
Template "01_One_Nav_Level" 1920x1080
   Gauge "gaugeDiagStateUpdate" at 566,2 size 50x50; CaptionText 'SIMATIC'
      on Change: "CheckDiagState"()
      ProcessValue <- "@DiagnosticsIndicatorTag"
   TextField "txtTitleBar" at 8,11 size 361x32; Text 'Application Name / Applikation / 江苏睿博环保再生胶系统'
   GraphicView "gfxNavigationIcon" at 1879,15 size 23x19; Picture "Hamburger_Icon"
   Button "btnNavigation" at 1862,0 size 56x48; TextOff 'Text'
      on Click: function_cf6f4242("GraphX_Slidein_Right", 1)
   TextField "模板_文本域_1" at 283,78 size 160x19; Text '全胎粉'
   TextField "txtTitleBar_1" at 12,1031 size 62x32; Text 'Application Name / Applikation / 冷水:'
   TextField "txtTitleBar_2" at 173,1031 size 62x32; Text 'Application Name / Applikation / 热水:'
   TextField "txtTitleBar_3" at 345,1031 size 62x32; Text 'Application Name / Applikation / 备料:'
   TextField "txtTitleBar_4" at 1752,1030 size 69x32; Text 'Application Name / Applikation / 数据库:'
   TextField "txtTitleBar_5" at 1587,1031 size 69x32; Text 'Application Name / Applikation / 云数据:'
   AlarmView "模板_报警视图_1" at 495,1024 size 1069x52
   IOField "I/O 域_58" at 1096,73 size 129x32; FormatPattern 999999.9; Unit  H
   IOField "I/O 域_59" at 1406,75 size 130x32; FormatPattern 99999999.9; Unit  Kg
   ScreenModuleView "HMI_Indicator_Square_1" at 1834,1033 size 28x28; ScreenModuleType ""
      Guid_{11997190-149293} <- "数据库字符串_Connect_CND"
      Guid_{11997190-149297} <- "数据库字符串_Query_Error"
      Guid_{11997190-149295} <- "数据库字符串_Query_Done"
   ScreenModuleView "HMI_Indicator_Square_2" at 1669,1033 size 28x28; ScreenModuleType ""
      Guid_{11997190-149295} <- "数据库字符串_Query_Done"
      Guid_{11997190-149293} <- "数据库字符串_Connect_CND"
      Guid_{11997190-149297} <- "数据库字符串_Query_Error"
   TextField "模板_文本域_2" at 77,80 size 73x19; Text '请选择'
   Button "btnStartscreen" at 1,2 size 411x45; TextOff 'Text'
      on Click: "ActivateStartScreen"()
   TextField "txtStateHeadline" at 75,55 size 123x23; Text 'State / Status / 运行配方'
   TextField "txtRecipeHeadline" at 281,55 size 154x23; Text 'Current Recipe / Rezeptur / 运行模式'
   TextField "txtOperatorHeadline" at 527,55 size 129x23; Text 'Operator / Bediener / 当前用户'
   IOField "ioOperator" at 527,72 size 126x30; FormatPattern ??????????????????
      ProcessValue <- "CurrentUserName"
   Button "btnState" at 202,56 size 40x40; TextOff '...'; PictureOff "More_Icon"
      on Click: "ShowRecipePopUp"()
   Button "btnRecipe" at 449,56 size 40x40; TextOff '...'; PictureOff "More_Icon"
   Rectangle "rectState" at 0,48 size 56x56
      Appearance <- "CurrentMachineState"
   GraphicIOField "gioDiagState" at 1874,60 size 32x32; PictureList "DiagState_3"
      ProcessValue <- "DiagState"
   Button "btnDiagState" at 1862,48 size 56x56; TextOff 'Text'
   Button "btnOperator" at 669,56 size 40x40; TextOff '...'; PictureOff "More_Icon"
      on Click: function_efd93a16("Template_Logon", 800, 300, -1, -1, 1)
   TextField "txtOperatorHeadline_1" at 768,55 size 129x23; Text 'Date and Time / Bediener / 当前时间'
   Button "btnOperator_1" at 995,56 size 40x40; TextOff '...'; PictureOff "More_Icon"
   DateTimeField "Template_Date/time field_1" at 768,72 size 208x30
   IOField "ioOperator_1" at 69,1033 size 99x30; FormatPattern 99.9; Unit m³/h
   IOField "ioOperator_2" at 230,1033 size 97x30; FormatPattern 99.9; Unit m³/h
   IOField "ioOperator_3" at 402,1033 size 72x30; FormatPattern 99.9; Unit %
   TextField "txtOperatorHeadline_2" at 1094,57 size 129x23; Text 'Date and Time / Bediener / 累计运行时间'
   Button "btnOperator_2" at 1321,58 size 40x40; TextOff '...'; PictureOff "More_Icon"
   TextField "txtOperatorHeadline_3" at 1403,58 size 129x23; Text 'Date and Time / Bediener / 累计产量'
   Button "btnOperator_3" at 1630,59 size 40x40; TextOff '...'; PictureOff "More_Icon"

PopupScreen "Template_Logon" 320x352
   on ClearScreen: ResetBit("PopUpBackground")
   on GenerateScreen: SetBit("PopUpBackground")
   TextField "Template_Text field_1" at 16,0 size 215x40; Text 'Login / 登录'
   Button "Button_2" at 16,240 size 288x40; TextOn 'LOGIN / ANMELDEN / 登录'; TextOff 'LOGIN / ANMELDEN / 登录'
      on Click: function_a9b89908("Password", "UserName"); function_efd93a16("Template_Logon", 0, 0, 0, -1, 1)
   IOField "I/O field_1" at 16,84 size 288x40; FormatPattern ??????????????????????????????
      ProcessValue <- "UserName"
   TextField "Text field_1" at 16,56 size 288x24; Text 'User Name / Name / 用户名'
   IOField "I/O field_2" at 16,168 size 288x40; FormatPattern ??????????????????????????????
      ProcessValue <- "Password"
   TextField "Text field_2" at 16,140 size 288x24; Text 'Password / Passwort / 密码'
   Button "Button_1" at 16,296 size 288x40; TextOn 'CLOSE / SCHLIESSEN / 取消'; TextOff 'CLOSE / SCHLIESSEN / 取消'
      on Click: function_efd93a16("Template_Logon", 0, 0, 0, -1, 1)
      on Press: function_b14e0dd5("ButtonDown", 0)
      Appearance <- "ButtonDown"

PopupScreen "Template_Logon_Logoff" 320x352
   on ClearScreen: ResetBit("PopUpBackground")
   on GenerateScreen: SetBit("PopUpBackground")
   TextField "Template_Text field_1" at 16,0 size 215x40; Text 'Login'
   Button "Button_2" at 16,240 size 136x40; TextOn 'LOG OFF / ABMELDEN'; TextOff 'LOG OFF / ABMELDEN'
      on Click: function_f23ef4c9()
   IOField "I/O field_1" at 16,84 size 288x40; FormatPattern ??????????????????????????????
      ProcessValue <- "UserName"
   TextField "Text field_1" at 16,56 size 288x24; Text 'User Name / Name'
   IOField "I/O field_2" at 16,168 size 288x40; FormatPattern ??????????????????????????????
      ProcessValue <- "Password"
   TextField "Text field_2" at 16,140 size 288x24; Text 'Password / Passwort'
   Button "Button_1" at 16,296 size 288x40; TextOn 'CLOSE / SCHLIESSEN'; TextOff 'CLOSE / SCHLIESSEN'
      on Click: function_efd93a16("Template_Logon_Logoff", 0, 0, 0, -1, 1)
      on Press: function_b14e0dd5("ButtonDown", 0)
      Appearance <- "ButtonDown"
   Button "Button_3" at 168,240 size 136x40; TextOn 'LOGIN / ANMELDEN'; TextOff 'LOGIN / ANMELDEN'
      on Click: function_a9b89908("Password", "UserName"); function_efd93a16("Template_Logon_Logoff", 0, 0, 0, -1, 1)

PopupScreen "Template_Operating_Mode" 424x360
   on ClearScreen: ResetBit("PopUpBackground")
   on GenerateScreen: SetBit("PopUpBackground")
   TextField "Template_Text field_1" at 14,0 size 336x40; Text 'Operating Mode / Betriebsmodus / 单螺杆操作'
   Button "Button_2" at 352,66 size 40x40; TextOff 'Text'; PictureOff "More_Icon"; PictureOn "More_Icon"
      on Click: function_efd93a16("Template_Operating_Mode", 0, 0, 0, -1, 1)
   Button "Button_3" at 352,130 size 40x40; TextOff 'Text'; PictureOff "More_Icon"; PictureOn "More_Icon"
      on Click: function_efd93a16("Template_Operating_Mode", 0, 0, 0, -1, 1)
   Button "Button_4" at 352,189 size 40x40; TextOff 'Text'; PictureOff "More_Icon"; PictureOn "More_Icon"
   Button "Button_1" at 352,254 size 40x40; TextOff 'Text'; PictureOff "More_Icon"; PictureOn "More_Icon"
   TextField "txtParameter7_3" at 32,63 size 163x24; Text 'Demo Mode / Current Mode / 演示模式'
   TextField "txtParameter7_5" at 31,89 size 319x24; Text 'Current Mode / 通过控制台仿真数据给触摸屏进行系统演示'
   TextField "txtParameter7_1" at 32,129 size 163x24; Text 'Test Mode / Current Mode / 测试模式'
   TextField "txtParameter7_2" at 31,155 size 319x24; Text 'Current Mode / 通过控制台仿真数据给触摸屏进行系统演示'

PopupScreen "Template_Recipe" 700x420
   on ClearScreen: ResetBit("PopUpBackground")
   on GenerateScreen: SetBit("PopUpBackground")
   TextField "Template_Text field_1" at 14,0 size 500x40; Text 'Recipe / Rezeptur'
   Button "Button_1" at 220,364 size 260x40; TextOn 'CLOSE / SCHLIESSEN'; TextOff 'CLOSE / SCHLIESSEN / 确定'
      on Click: function_efd93a16("Template_Recipe", 0, 0, 0, -1, 1)
      on Press: function_b14e0dd5("ButtonDown", 0)
      Appearance <- "ButtonDown"

PopupScreen "OptionPanel_4_Buttons_1" 390x648
   Button "btnCloseOptionPanel" at 0,0 size 40x648; TextOff 'CLOSE'; PictureOff "Jog_Forward"
      on Press: function_efd93a16("OptionPanel_4_Buttons_1", 0, 0, 0, 2, 2)
   TextField "txtOptionPanel" at 108,16 size 260x40; Text 'Option Panel Title / Titel Option Panel'
   Button "btnOption1" at 80,72 size 240x40; TextOff 'Option 1 / Move to Home Position'
   Button "btnOption2" at 80,128 size 240x40; TextOff 'Option 2 / Move to Home Position'
   Button "btnOption3" at 80,184 size 240x40; TextOff 'Option 3 / RESET'
   Button "btnOption4" at 80,240 size 240x40; TextOff 'Option 4 / RESET'
   GraphicView "gvOptionPanel" at 80,30 size 18x12; Picture "ManFunctions_Off"

PopupScreen "OptionPanel_4_Buttons" 390x648
   Button "btnCloseOptionPanel" at 0,0 size 40x648; TextOff 'CLOSE'; PictureOff "Jog_Forward"
      on Press: function_efd93a16("OptionPanel_4_Buttons", 0, 0, 0, 2, 2)
   TextField "txtOptionPanel" at 108,16 size 260x40; Text 'Option Panel Title / Titel Option Panel'
   Button "btnOption1" at 80,72 size 240x40; TextOff 'Option 1 / Move to Home Position'
   Button "btnOption2" at 80,128 size 240x40; TextOff 'Option 2 / Move to Home Position'
   Button "btnOption3" at 80,184 size 240x40; TextOff 'Option 3 / RESET'
   Button "btnOption4" at 80,240 size 240x40; TextOff 'Option 4 / RESET'
   GraphicView "gvOptionPanel" at 80,30 size 18x12; Picture "ManFunctions_Off"

PopupScreen "OptionPanel_4_Large_Buttons" 390x648
   Button "btnCloseOptionPanel" at 0,0 size 40x648; TextOff 'CLOSE'; PictureOff "Jog_Forward"
      on Press: function_efd93a16("OptionPanel_4_Large_Buttons", 0, 0, 0, 2, 2)
   TextField "txtOptionPanel" at 108,16 size 260x40; Text 'Option Panel Title / Titel Option Panel'
   GraphicView "gvOptionPanel" at 80,30 size 18x12; Picture "ManFunctions_Off"
   Button "btnOption1" at 80,72 size 112x96; TextOff 'Option 1 / Move to Home Position'
   Button "btnOption2" at 208,72 size 112x96; TextOff 'Option 2 / Move to Home Position'
   Button "btnOption3" at 80,184 size 112x96; TextOff 'Option 3 / Move to Home Position'
   Button "btnOption4" at 208,184 size 112x96; TextOff 'Option 4 / Move to Home Position'

PopupScreen "OptionPanel_8_Buttons" 390x648
   Button "btnCloseOptionPanel" at 0,0 size 40x648; TextOff 'CLOSE'; PictureOff "Jog_Forward"
      on Press: function_efd93a16("OptionPanel_8_Buttons", 0, 0, 0, 2, 2)
   TextField "txtOptionPanel" at 108,16 size 260x40; Text 'Option Panel Title / Titel Option Panel'
   GraphicView "gvOptionPanel" at 80,30 size 18x12; Picture "ManFunctions_Off"
   Button "btnOption1" at 80,72 size 112x40; TextOff 'Option 1 / Move to Home Position'
   Button "btnOption2" at 208,72 size 112x40; TextOff 'Option 2 / Move to Home Position'
   Button "btnOption3" at 80,128 size 112x40; TextOff 'Option 3 / Move to Home Position'
   Button "btnOption4" at 208,128 size 112x40; TextOff 'Option 4 / Move to Home Position'
   Button "btnOption5" at 80,184 size 112x40; TextOff 'Option 5 / Move to Home Position'
   Button "btnOption6" at 208,184 size 112x40; TextOff 'Option 6 / Move to Home Position'
   Button "btnOption7" at 80,240 size 112x40; TextOff 'Option 7 / Move to Home Position'
   Button "btnOption8" at 208,240 size 112x40; TextOff 'Option 8 / Move to Home Position'

PopupScreen "OptionPanel_8_Large_Buttons" 390x648
   Button "btnCloseOptionPanel" at 0,0 size 40x648; TextOff 'CLOSE'; PictureOff "Jog_Forward"
      on Press: function_efd93a16("OptionPanel_8_Large_Buttons", 0, 0, 0, 2, 2)
   TextField "txtOptionPanel" at 108,16 size 260x40; Text 'Option Panel Title / Titel Option Panel'
   GraphicView "gvOptionPanel" at 80,30 size 18x12; Picture "ManFunctions_Off"
   Button "btnOption1" at 80,72 size 112x96; TextOff 'Option 1 / Move to Home Position'
   Button "btnOption2" at 208,72 size 112x96; TextOff 'Option 2 / Move to Home Position'
   Button "btnOption3" at 80,184 size 112x96; TextOff 'Option 3 / Move to Home Position'
   Button "btnOption4" at 208,184 size 112x96; TextOff 'Option 4 / Move to Home Position'
   Button "btnOption5" at 80,296 size 112x96; TextOff 'Option 1 / Option 5 / Move to Home Position'
   Button "btnOption6" at 208,296 size 112x96; TextOff 'Option 2 / Option 6 / Move to Home Position'
   Button "btnOption7" at 80,408 size 112x96; TextOff 'Option 3 / Option 7 / Move to Home Position'
   Button "btnOption8" at 208,408 size 112x96; TextOff 'Option 4 / Option 8 / Move to Home Position'

PopupScreen "BM00_Operating" 424x360
   on ClearScreen: ResetBit("PopUpBackground")
   on GenerateScreen: SetBit("PopUpBackground")
   TextField "Template_Text field_1" at 14,0 size 336x40; Text 'Operating Mode / Betriebsmodus / BM00控制'
   Button "Button_2" at 62,310 size 288x40; TextOn 'LOGIN / ANMELDEN / 登录'; TextOff 'LOGIN / ANMELDEN / 确定'
      on Click: function_efd93a16("BM00_Operating", 0, 0, 0, -1, 1)

SlideinScreen "GraphX_Slidein_Right" 250x1080
   Button "Button_1" at 9,164 size 220x60; TextOn 'MainView / Menu Item 1 / 主界面'; TextOff 'MainView / Menu Item 1 / 数据看板'
      on Click: SetTag("MainNavigationState", 1); ActivateScreen("监控主画面", 0)
      Appearance <- "MainNavigationState"
   Button "Button_2" at 9,226 size 220x60; TextOn 'S.W.Pump / Menu Item 2 / 海水泵'; TextOff 'S.W.Pump / Menu Item 2 / 精炼监控'
      on Click: SetTag("MainNavigationState", 2)
      Appearance <- "MainNavigationState"
   Button "Button_3" at 9,287 size 220x60; TextOn 'Pump(S) / Menu Item 3 / 泵组'; TextOff 'Pump(S) / Menu Item 3 / 水 系 统'
      on Click: SetTag("MainNavigationState", 3)
      Appearance <- "MainNavigationState"
   Rectangle "Rectangle_1" at 223,164 size 6x60
      Visibility <- "MainNavigationState"
   Rectangle "Rectangle_2" at 223,226 size 6x60
      Visibility <- "MainNavigationState"
   Rectangle "Rectangle_3" at 223,287 size 6x60
      Visibility <- "MainNavigationState"
   Button "Button_4" at 9,348 size 220x60; TextOn 'Valve(S) / Menu Item 4 / 阀组'; TextOff 'Valve(S) / Menu Item 4 / 报表统计'
      on Click: SetTag("MainNavigationState", 4)
      Appearance <- "MainNavigationState"
   Rectangle "Rectangle_4" at 223,348 size 6x60
      Visibility <- "MainNavigationState"
   Button "Button_5" at 9,410 size 220x60; TextOn 'Menu Item 4 / 烟气监测'; TextOff 'Settings / Menu Item 4 / 工艺设置'
      on Click: SetTag("MainNavigationState", 5)
      Appearance <- "MainNavigationState"
   Rectangle "Rectangle_5" at 223,410 size 6x60
      Visibility <- "MainNavigationState"
   Button "Button_6" at 9,472 size 220x60; TextOn 'Menu Item 4 / 水质监测'; TextOff 'Settings / Menu Item 4 / 系统设置'
      on Click: SetTag("MainNavigationState", 6)
      Appearance <- "MainNavigationState"
   Rectangle "Rectangle_6" at 223,472 size 6x60
      Visibility <- "MainNavigationState"
   Button "Button_7" at 9,534 size 220x60; TextOn 'Other(S) / Menu Item 4 / 其他'; TextOff 'Other(S) / Menu Item 4 / 其他'
      on Click: SetTag("MainNavigationState", 7)
      Appearance <- "MainNavigationState"
   Rectangle "Rectangle_7" at 223,534 size 6x60
      Visibility <- "MainNavigationState"
   Button "Button_8" at 9,596 size 220x60; TextOn 'Spare / Menu Item 4 / 备用'; TextOff 'Spare / Menu Item 4 / 报警列表'
      on Click: SetTag("MainNavigationState", 8)
      Appearance <- "MainNavigationState"
   Rectangle "Rectangle_8" at 223,596 size 6x60
      Visibility <- "MainNavigationState"
   Button "Button_9" at 9,658 size 220x60; TextOn 'Settings / Menu Item 4 / 设置'; TextOff 'Settings / Menu Item 4 / 帮助'
      on Click: SetTag("MainNavigationState", 9)
      Appearance <- "MainNavigationState"
   Rectangle "Rectangle_9" at 223,658 size 6x60
      Visibility <- "MainNavigationState"

screen "监控主画面" 1920x1080, template "01_One_Nav_Level"
   ScreenModuleView "精炼机面板_1" at 17,115 size 338x480; ScreenModuleType ""
      Guid_{11997190-15377} <- "数据库字符串_Upload{11}"
   ScreenModuleView "精炼机面板_2" at 397,115 size 338x480; ScreenModuleType ""; Guid_{11997190-15477} 'N12号精炼机'
      Guid_{11997190-15377} <- "数据库字符串_Upload{12}"
   ScreenModuleView "精炼机面板_3" at 781,115 size 338x480; ScreenModuleType ""; Guid_{11997190-15477} 'N13号精炼机'
      Guid_{11997190-15377} <- "数据库字符串_Upload{13}"
   ScreenModuleView "精炼机面板_4" at 1160,115 size 338x480; ScreenModuleType ""; Guid_{11997190-15477} 'N14号精炼机'
      Guid_{11997190-15377} <- "数据库字符串_Upload{14}"
   ScreenModuleView "精炼机面板_5" at 1536,115 size 338x480; ScreenModuleType ""; Guid_{11997190-15477} 'N15号精炼机'
      Guid_{11997190-15377} <- "数据库字符串_Upload{15}"
   TextField "文本域_1" at 32,611 size 65x23; Text '环境温度'
   IOField "I/O 域_1" at 32,631 size 234x71; FormatPattern 99.9
      ProcessValue <- "通用数据采集_环境温度"
   TextField "文本域_2" at 261,678 size 20x23; Text '℃'
   TextField "文本域_3" at 32,741 size 65x23; Text '环境湿度'
   IOField "I/O 域_2" at 32,763 size 228x71; FormatPattern 99.9
      ProcessValue <- "通用数据采集_环境湿度"
   TextField "文本域_4" at 259,810 size 41x23; Text '%RH'
   TextField "文本域_5" at 33,872 size 50x23; Text '循环水'
   IOField "I/O 域_3" at 33,894 size 224x71; FormatPattern 99.9
   TextField "文本域_6" at 260,941 size 20x23; Text '℃'
   TextField "文本域_7" at 1552,614 size 96x23; Text 'N21累计产量'
   IOField "I/O 域_4" at 1551,634 size 313x71; FormatPattern 9999999999
      ProcessValue <- "精炼机数据转存_N21卷片机累计重量"
   TextField "文本域_8" at 1844,684 size 25x23; Text 'Kg'
   TextField "文本域_9" at 1556,745 size 96x23; Text 'N22累计产量'
   IOField "I/O 域_5" at 1552,765 size 313x71; FormatPattern 9999999999
      ProcessValue <- "精炼机数据转存_N22卷片机累计重量"
   TextField "文本域_10" at 1849,814 size 25x23; Text 'Kg'

VB script "MainEntry"
   bec8f1e5-2ab1-45f6-ad91-1d37c469eb91 监控主画面, 0

VB script "ActivateAlarmControlScreen"
   bec8f1e5-2ab1-45f6-ad91-1d37c469eb91 20_Messages,0

VB script "ActivateStartScreen"
   HmiRuntime.BaseScreenName = SmartTags("StartScreenName")

VB script "CheckCurrentLanguage"
   If HmiRuntime.Language = 1031 Then 'German
   	SmartTags("CurrentLanguage") = 0
   	ElseIf HmiRuntime.Language = 1033 Then 'English US
   	SmartTags("CurrentLanguage") = 1
   End If
   
   	

VB script "CheckCurrentUserName"
   If SmartTags("CurrentUserName") = "" Or SmartTags("CurrentUserName") = "User Name" Or SmartTags("CurrentUserName") = "Benutzer" Then
     
     If HmiRuntime.Language = 1031 Then 'Germany
       SmartTags("CurrentUserName") = "Benutzer"
       
     ElseIf HmiRuntime.Language = 1033 Then 'English US
       SmartTags("CurrentUserName") = "User Name"
     End If
     
     SmartTags("UserIsLoggedIn") = False
   Else
     If SmartTags("CurrentUserName") <> "User Name" And SmartTags("CurrentUserName") <> "Benutzer" Then
       SmartTags("UserIsLoggedIn") = True  
     End If
   End If

VB script "CheckDiagState"
   If SmartTags("@DiagnosticsIndicatorTag") = 1 Then
   	SmartTags("DiagState") = 1
   Else
   	SmartTags("DiagState") = 0
   End If

VB script "GetStartScreenName"
   SmartTags("StartScreenName") = HmiRuntime.BaseScreenName

VB script "ShowLoginPopUp"
   efd93a16-2665-4b85-bcb9-25eddcb7b6f4 Template_Logon_Logoff,480,110,$3$hmiOn$,$3$hmiAnimationOff$,$3$hmiFast$

VB script "ShowOperatingModePopUp"
   efd93a16-2665-4b85-bcb9-25eddcb7b6f4 Template_Operating_Mode,800,300,$3$hmiOn$,$3$hmiAnimationOff$,$3$hmiFast$

VB script "ShowOptionPanelPopUp"
   efd93a16-2665-4b85-bcb9-25eddcb7b6f4 OptionPanel_4_Buttons, 890, 110, $3$hmiOn$, $3$hmiRight$, $3$hmiFast$

VB script "ShowRecipePopUp"
   efd93a16-2665-4b85-bcb9-25eddcb7b6f4 Template_Recipe,290,110,$3$hmiOn$,$3$hmiAnimationOff$,$3$hmiFast$

VB script "ShowSimAnalog"
   efd93a16-2665-4b85-bcb9-25eddcb7b6f4 Template_Sim_Analog_Set,800,300,$3$hmiOn$,$3$hmiAnimationOff$,$3$hmiFast$

VB script "ShowSimValve"
   efd93a16-2665-4b85-bcb9-25eddcb7b6f4 Template_Sim_Valve_Set,800,300,$3$hmiOn$,$3$hmiAnimationOff$,$3$hmiFast$

VB script "ShowSimProfidrive"
   efd93a16-2665-4b85-bcb9-25eddcb7b6f4 Template_Sim_Profidrive,800,300,$3$hmiOn$,$3$hmiAnimationOff$,$3$hmiFast$

VB script "ShowSimME"
   efd93a16-2665-4b85-bcb9-25eddcb7b6f4 Template_Sim_ME_Set,800,300,$3$hmiOn$,$3$hmiAnimationOff$,$3$hmiFast$
*)

(* ===== HMI "HMI_RT_1" =====

ScreenModuleEditorView "HMI_Indicator_Square" 640x480
   Rectangle "Ready" at 10,10 size 116x93
      Visibility <- "备妥"
   Rectangle "Running" at 10,10 size 116x93
      Visibility <- "运行"
   Rectangle "Fault" at 10,10 size 116x93
      Visibility <- "故障"
*)

(* ===== HMI "HMI_RT_1" =====
system functions are stored by id; their names below are inferred from use

text list "按钮名称": 0 'ON'; 1 'OFF'

ScreenModuleEditorView "OnKey" 640x480
   Rectangle "矩形_1" at 13,9 size 67x29
      Appearance <- "参数.Fault"
   TextField "文本域_1" at 19,12 size 53x23; Text 'FAULT'
   Button "按钮_2" at 9,8 size 74x31; TextOff 'Text'; TextList "按钮名称"
      on Click: SetTag("参数.Stop", "参数.Running"); InvertBit("参数.Running"); SetTag("参数.Start", "参数.Running")
      Visibility <- "参数.Ready"
      ProcessValue <- "参数.Running"
      Appearance <- "参数.Running"
*)

(* ===== HMI "HMI_RT_1" =====

HMI tags "默认变量表"
   "Step" : Int, internal

ScreenModuleEditorView "流程步骤控制" 640x480
   Button "按钮_1" at 10,10 size 38x41; TextOff '1'
   Button "按钮_2" at 51,10 size 294x41; TextOff '检测混料系统备妥'
      Appearance <- "变量.StepRuning"
   Button "按钮_3" at 347,10 size 98x41; TextOff 'OK'
      Appearance <- "变量.StepOK"
   Button "按钮_4" at 347,10 size 98x41; TextOff 'NOK'
      Visibility <- "变量.StepNok"

VB script "FaceplateScript_1"
   '提示：
   ' 1. 使用 <CTRL+SPACE> 或 <CTRL+I> 快捷键打开含所有对象和函数的列表
   ' 2. 使用 HMI Runtime 对象写入代码。
   '  示例：HmiRuntime.Screens("Screen_1")。
   ' 3. 使用 <CTRL+J> 快捷键创建对象引用。
   '从此位置起写入代码：
*)

(* ===== HMI "HMI_RT_1" =====

ScreenModuleEditorView "HMI_Indicator_Square" 640x480
   Rectangle "Ready" at 10,10 size 116x93
      Visibility <- "备妥"
   Rectangle "Running" at 10,10 size 116x93
      Visibility <- "运行"
   Rectangle "Fault" at 10,10 size 116x93
      Visibility <- "故障"
*)

(* ===== HMI "HMI_RT_1" =====

ScreenModuleEditorView "精炼机面板" 640x480
   TextField "Template_Text field_1" at 10,10 size 336x40; Text 'Operating Mode / Betriebsmodus / NO.11'
*)

(* ===== HMI "HMI_RT_1" =====

ScreenModuleEditorView "精炼机面板" 380x480
   Rectangle "备妥矩形" at 1,1 size 377x48
      Visibility <- "数据变量.开关量汇总"
   Rectangle "运行矩形" at 1,1 size 377x48
      Visibility <- "数据变量.开关量汇总"
   Rectangle "故障矩形" at 1,1 size 377x48
      Visibility <- "数据变量.开关量汇总"
   TextField "设备名称" at 8,7 size 145x35; Text 'N11号精炼机'
   IOField "I/O 域_1" at 8,72 size 154x80; FormatPattern 999
   IOField "I/O 域_2" at 8,170 size 160x80; FormatPattern 99.9
   TextField "文本域_2" at 163,221 size 28x26; Text 'HZ'
   TextField "文本域_3" at 163,135 size 17x26; Text 'A'
   TextField "文本域_4" at 9,49 size 37x26; Text '电流'
   TextField "文本域_5" at 9,148 size 37x26; Text '频率'
   IOField "I/O 域_3" at 199,69 size 154x80; FormatPattern 999
   TextField "文本域_1" at 358,132 size 20x26; Text '%'
   TextField "文本域_6" at 200,46 size 37x26; Text '功率'
   IOField "I/O 域_4" at 202,172 size 154x80; FormatPattern 999
   TextField "文本域_7" at 356,235 size 21x26; Text '℃'
   TextField "文本域_8" at 203,149 size 37x26; Text '胶温'
*)

(* ===== HMI "HMI_RT_1" =====

ScreenModuleEditorView "精炼机面板" 380x480
   Rectangle "备妥矩形" at 1,1 size 377x48
      Visibility <- "数据变量.开关量汇总"
   Rectangle "运行矩形" at 1,1 size 377x48
      Visibility <- "数据变量.开关量汇总"
   Rectangle "故障矩形" at 1,1 size 377x48
      Visibility <- "数据变量.开关量汇总"
   TextField "设备名称" at 8,7 size 145x35; Text 'N11号精炼机'
   IOField "I/O 域_1" at 8,72 size 154x80; FormatPattern 999
      ProcessValue <- "数据变量.滚筒电机电流"
   IOField "I/O 域_2" at 8,170 size 160x80; FormatPattern 99.9
      ProcessValue <- "数据变量.滚筒电机频率"
   TextField "文本域_2" at 163,221 size 28x26; Text 'HZ'
   TextField "文本域_3" at 163,135 size 17x26; Text 'A'
   TextField "文本域_4" at 9,49 size 37x26; Text '电流'
   TextField "文本域_5" at 9,148 size 37x26; Text '频率'
   IOField "I/O 域_3" at 199,69 size 154x80; FormatPattern 999
      ProcessValue <- "数据变量.滚筒电机功率"
   TextField "文本域_1" at 358,132 size 20x26; Text '%'
   TextField "文本域_6" at 200,46 size 37x26; Text '功率'
   IOField "I/O 域_4" at 202,172 size 154x80; FormatPattern 999
      ProcessValue <- "数据变量.胶温"
   TextField "文本域_7" at 356,235 size 21x26; Text '℃'
   TextField "文本域_8" at 203,149 size 37x26; Text '胶温'
   TextField "文本域_9" at 8,450 size 35x23; Text '计时:'
   TextField "文本域_10" at 177,450 size 35x23; Text '电能:'
   IOField "I/O 域_5" at 43,454 size 90x17; FormatPattern 9999999999
      ProcessValue <- "数据变量.滚筒电机计时"
   TextField "文本域_11" at 142,451 size 13x23; Text 'S'
   IOField "I/O 域_6" at 212,454 size 90x17; FormatPattern 9999999999
      ProcessValue <- "数据变量.滚筒电机电度"
   TextField "文本域_12" at 308,451 size 39x23; Text 'KWH'
   TextField "文本域_13" at 17,268 size 87x23; Text '左前滚筒轴温:'
   IOField "I/O 域_7" at 50,286 size 82x43; FormatPattern 999.9
      ProcessValue <- "数据变量.左前辊温度"
   TextField "文本域_14" at 163,298 size 18x23; Text '℃'
   TextField "文本域_15" at 204,268 size 87x23; Text '右前滚筒轴温:'
   IOField "I/O 域_8" at 237,286 size 82x43; FormatPattern 999.9
      ProcessValue <- "数据变量.右前辊温度"
   TextField "文本域_16" at 350,298 size 18x23; Text '℃'
   TextField "文本域_17" at 16,319 size 87x23; Text '左后滚筒轴温:'
   IOField "I/O 域_9" at 49,337 size 82x43; FormatPattern 999.9
      ProcessValue <- "数据变量.左后辊温度"
   TextField "文本域_18" at 162,349 size 18x23; Text '℃'
   TextField "文本域_19" at 204,320 size 87x23; Text '右后滚筒轴温:'
   IOField "I/O 域_10" at 237,338 size 82x43; FormatPattern 999.9
      ProcessValue <- "数据变量.右后辊温度"
   TextField "文本域_20" at 350,350 size 18x23; Text '℃'
   TextField "文本域_21" at 17,374 size 83x23; Text '左滚筒间隙值'
   IOField "I/O 域_11" at 50,392 size 82x43; FormatPattern 9999
      ProcessValue <- "数据变量.左间隙"
   TextField "文本域_22" at 163,404 size 18x23; Text '丝'
   TextField "文本域_23" at 205,377 size 87x23; Text '右滚筒间隙值:'
   IOField "I/O 域_12" at 238,391 size 82x43; FormatPattern 9999
      ProcessValue <- "数据变量.右间隙"
   TextField "文本域_24" at 351,403 size 18x23; Text '丝'
   IOField "I/O 域_13" at 204,6 size 164x45; FormatPattern ????
      ProcessValue <- "数据变量.当前人员编号"
*)

(* ===== HMI "HMI_RT_1" =====

ScreenModuleEditorView "精炼机面板" 380x480
   Rectangle "备妥矩形" at 1,1 size 377x48
      Visibility <- "数据变量.开关量汇总"
   Rectangle "运行矩形" at 1,1 size 377x48
      Visibility <- "数据变量.开关量汇总"
   Rectangle "故障矩形" at 1,1 size 377x48
      Visibility <- "数据变量.开关量汇总"
   TextField "设备名称" at 8,7 size 145x35; Text 'N11号精炼机'
   IOField "I/O 域_1" at 8,72 size 154x80; FormatPattern 999
      ProcessValue <- "数据变量.滚筒电机电流"
   IOField "I/O 域_2" at 8,170 size 160x80; FormatPattern 99.9
      ProcessValue <- "数据变量.滚筒电机频率"
   TextField "文本域_2" at 163,221 size 28x26; Text 'HZ'
   TextField "文本域_3" at 163,135 size 17x26; Text 'A'
   TextField "文本域_4" at 9,49 size 37x26; Text '电流'
   TextField "文本域_5" at 9,148 size 37x26; Text '频率'
   IOField "I/O 域_3" at 199,69 size 154x80; FormatPattern 999
      ProcessValue <- "数据变量.滚筒电机功率"
   TextField "文本域_1" at 358,132 size 20x26; Text '%'
   TextField "文本域_6" at 200,46 size 37x26; Text '功率'
   IOField "I/O 域_4" at 202,172 size 154x80; FormatPattern 999
      ProcessValue <- "数据变量.胶温"
   TextField "文本域_7" at 356,235 size 21x26; Text '℃'
   TextField "文本域_8" at 203,149 size 37x26; Text '胶温'
   TextField "文本域_9" at 8,450 size 35x23; Text '计时:'
   TextField "文本域_10" at 177,450 size 35x23; Text '电能:'
   IOField "I/O 域_5" at 43,454 size 90x17; FormatPattern 9999999999
      ProcessValue <- "数据变量.滚筒电机计时"
   TextField "文本域_11" at 142,451 size 13x23; Text 'S'
   IOField "I/O 域_6" at 212,454 size 90x17; FormatPattern 9999999999
      ProcessValue <- "数据变量.滚筒电机电度"
   TextField "文本域_12" at 308,451 size 39x23; Text 'KWH'
   TextField "文本域_13" at 17,268 size 87x23; Text '左前滚筒轴温:'
   IOField "I/O 域_7" at 50,286 size 82x43; FormatPattern 999.9
      ProcessValue <- "数据变量.左前辊温度"
   TextField "文本域_14" at 163,298 size 18x23; Text '℃'
   TextField "文本域_15" at 204,268 size 87x23; Text '右前滚筒轴温:'
   IOField "I/O 域_8" at 237,286 size 82x43; FormatPattern 999.9
      ProcessValue <- "数据变量.右前辊温度"
   TextField "文本域_16" at 350,298 size 18x23; Text '℃'
   TextField "文本域_17" at 16,319 size 87x23; Text '左后滚筒轴温:'
   IOField "I/O 域_9" at 49,337 size 82x43; FormatPattern 999.9
      ProcessValue <- "数据变量.左后辊温度"
   TextField "文本域_18" at 162,349 size 18x23; Text '℃'
   TextField "文本域_19" at 204,320 size 87x23; Text '右后滚筒轴温:'
   IOField "I/O 域_10" at 237,338 size 82x43; FormatPattern 999.9
      ProcessValue <- "数据变量.右后辊温度"
   TextField "文本域_20" at 350,350 size 18x23; Text '℃'
   TextField "文本域_21" at 17,374 size 83x23; Text '左滚筒间隙值'
   IOField "I/O 域_11" at 50,392 size 82x43; FormatPattern 9999
      ProcessValue <- "数据变量.左间隙"
   TextField "文本域_22" at 163,404 size 18x23; Text '丝'
   TextField "文本域_23" at 205,377 size 87x23; Text '右滚筒间隙值:'
   IOField "I/O 域_12" at 238,391 size 82x43; FormatPattern 9999
      ProcessValue <- "数据变量.右间隙"
   TextField "文本域_24" at 351,403 size 18x23; Text '丝'
   IOField "I/O 域_13" at 204,6 size 164x45; FormatPattern ????
      ProcessValue <- "数据变量.当前人员编号"
*)

(* ===== HMI "HMI_RT_1" =====

ScreenModuleEditorView "精炼机面板" 380x480
   Rectangle "备妥矩形" at 1,1 size 377x48
      Visibility <- "数据变量.开关量汇总"
   Rectangle "运行矩形" at 1,1 size 377x48
      Visibility <- "数据变量.开关量汇总"
   Rectangle "故障矩形" at 1,1 size 377x48
      Visibility <- "数据变量.开关量汇总"
   TextField "设备名称" at 8,7 size 145x35; Text 'N11号精炼机'
   IOField "I/O 域_1" at 8,72 size 154x80; FormatPattern 999
      ProcessValue <- "数据变量.滚筒电机电流"
   IOField "I/O 域_2" at 8,170 size 160x80; FormatPattern 99.9
      ProcessValue <- "数据变量.滚筒电机频率"
   TextField "文本域_2" at 163,221 size 28x26; Text 'HZ'
   TextField "文本域_3" at 163,135 size 17x26; Text 'A'
   TextField "文本域_4" at 9,49 size 37x26; Text '电流'
   TextField "文本域_5" at 9,148 size 37x26; Text '频率'
   IOField "I/O 域_3" at 199,69 size 154x80; FormatPattern 999
      ProcessValue <- "数据变量.滚筒电机功率"
   TextField "文本域_1" at 358,132 size 20x26; Text '%'
   TextField "文本域_6" at 200,46 size 37x26; Text '功率'
   IOField "I/O 域_4" at 202,172 size 154x80; FormatPattern 999
      ProcessValue <- "数据变量.胶温"
   TextField "文本域_7" at 356,235 size 21x26; Text '℃'
   TextField "文本域_8" at 203,149 size 37x26; Text '胶温'
   TextField "文本域_9" at 8,450 size 35x23; Text '计时:'
   TextField "文本域_10" at 177,450 size 35x23; Text '电能:'
   IOField "I/O 域_5" at 43,454 size 90x17; FormatPattern 9999999999
      ProcessValue <- "数据变量.滚筒电机计时"
   TextField "文本域_11" at 142,451 size 13x23; Text 'S'
   IOField "I/O 域_6" at 212,454 size 90x17; FormatPattern 9999999999
      ProcessValue <- "数据变量.滚筒电机电度"
   TextField "文本域_12" at 308,451 size 39x23; Text 'KWH'
   TextField "文本域_13" at 17,268 size 87x23; Text '左前滚筒轴温:'
   IOField "I/O 域_7" at 50,286 size 82x43; FormatPattern 999.9
      ProcessValue <- "数据变量.左前辊温度"
   TextField "文本域_14" at 163,298 size 18x23; Text '℃'
   TextField "文本域_15" at 204,268 size 87x23; Text '右前滚筒轴温:'
   IOField "I/O 域_8" at 237,286 size 82x43; FormatPattern 999.9
      ProcessValue <- "数据变量.右前辊温度"
   TextField "文本域_16" at 350,298 size 18x23; Text '℃'
   TextField "文本域_17" at 16,328 size 87x23; Text '左后滚筒轴温:'
   IOField "I/O 域_9" at 49,346 size 82x43; FormatPattern 999.9
      ProcessValue <- "数据变量.左后辊温度"
   TextField "文本域_18" at 162,358 size 18x23; Text '℃'
   TextField "文本域_19" at 204,329 size 87x23; Text '右后滚筒轴温:'
   IOField "I/O 域_10" at 237,347 size 82x43; FormatPattern 999.9
      ProcessValue <- "数据变量.右后辊温度"
   TextField "文本域_20" at 350,359 size 18x23; Text '℃'
   TextField "文本域_21" at 17,392 size 83x23; Text '左滚筒间隙值'
   IOField "I/O 域_11" at 50,410 size 82x43; FormatPattern 9999
      ProcessValue <- "数据变量.左间隙"
   TextField "文本域_22" at 163,422 size 18x23; Text '丝'
   TextField "文本域_23" at 205,393 size 87x23; Text '右滚筒间隙值:'
   IOField "I/O 域_12" at 238,410 size 82x43; FormatPattern 9999
      ProcessValue <- "数据变量.右间隙"
   TextField "文本域_24" at 351,422 size 18x23; Text '丝'
   IOField "I/O 域_13" at 204,6 size 164x45; FormatPattern ????
      ProcessValue <- "数据变量.当前人员编号"
*)

(* ===== HMI "HMI_RT_1" =====

ScreenModuleEditorView "精炼机面板" 338x480
   Rectangle "备妥矩形" at 1,1 size 339x48
      Visibility <- "数据变量.开关量汇总"
   Rectangle "运行矩形" at 1,1 size 337x48
      Visibility <- "数据变量.开关量汇总"
   Rectangle "故障矩形" at 1,1 size 338x48
      Visibility <- "数据变量.开关量汇总"
   TextField "设备名称" at 8,11 size 107x28; Text 'N11号精炼机'
   IOField "I/O 域_1" at 8,72 size 154x80; FormatPattern 999
      ProcessValue <- "数据变量.滚筒电机电流"
   IOField "I/O 域_2" at 8,170 size 160x80; FormatPattern 99.9
      ProcessValue <- "数据变量.滚筒电机频率"
   TextField "文本域_2" at 118,218 size 28x26; Text 'HZ'
   TextField "文本域_3" at 118,132 size 17x26; Text 'A'
   TextField "文本域_4" at 9,49 size 37x26; Text '电流'
   TextField "文本域_5" at 9,148 size 37x26; Text '频率'
   IOField "I/O 域_3" at 199,69 size 154x80; FormatPattern 999
      ProcessValue <- "数据变量.滚筒电机功率"
   TextField "文本域_1" at 311,136 size 20x26; Text '%'
   TextField "文本域_6" at 200,46 size 37x26; Text '功率'
   IOField "I/O 域_4" at 202,172 size 154x80; FormatPattern 999
      ProcessValue <- "数据变量.胶温"
   TextField "文本域_7" at 309,218 size 21x26; Text '℃'
   TextField "文本域_8" at 203,149 size 37x26; Text '胶温'
   TextField "文本域_9" at 3,450 size 35x23; Text '计时:'
   TextField "文本域_10" at 158,450 size 35x23; Text '电能:'
   IOField "I/O 域_5" at 38,454 size 90x17; FormatPattern 9999999999
      ProcessValue <- "数据变量.滚筒电机计时"
   TextField "文本域_11" at 137,451 size 13x23; Text 'S'
   IOField "I/O 域_6" at 193,454 size 90x17; FormatPattern 9999999999
      ProcessValue <- "数据变量.滚筒电机电度"
   TextField "文本域_12" at 289,451 size 39x23; Text 'KWH'
   TextField "文本域_13" at 17,268 size 87x23; Text '左前滚筒轴温:'
   IOField "I/O 域_7" at 17,285 size 82x43; FormatPattern 999.9
      ProcessValue <- "数据变量.左前辊温度"
   TextField "文本域_14" at 109,297 size 18x23; Text '℃'
   TextField "文本域_15" at 204,268 size 87x23; Text '右前滚筒轴温:'
   IOField "I/O 域_8" at 201,284 size 82x43; FormatPattern 999.9
      ProcessValue <- "数据变量.右前辊温度"
   TextField "文本域_16" at 308,296 size 18x23; Text '℃'
   TextField "文本域_17" at 16,328 size 87x23; Text '左后滚筒轴温:'
   IOField "I/O 域_9" at 16,346 size 82x43; FormatPattern 999.9
      ProcessValue <- "数据变量.左后辊温度"
   TextField "文本域_18" at 108,357 size 18x23; Text '℃'
   TextField "文本域_19" at 204,329 size 87x23; Text '右后滚筒轴温:'
   IOField "I/O 域_10" at 201,345 size 82x43; FormatPattern 999.9
      ProcessValue <- "数据变量.右后辊温度"
   TextField "文本域_20" at 308,357 size 18x23; Text '℃'
   TextField "文本域_21" at 17,392 size 83x23; Text '左滚筒间隙值'
   IOField "I/O 域_11" at 12,408 size 82x43; FormatPattern 9999
      ProcessValue <- "数据变量.左间隙"
   TextField "文本域_22" at 109,421 size 18x23; Text '丝'
   TextField "文本域_23" at 205,393 size 87x23; Text '右滚筒间隙值:'
   IOField "I/O 域_12" at 200,408 size 82x43; FormatPattern 9999
      ProcessValue <- "数据变量.右间隙"
   TextField "文本域_24" at 309,420 size 18x23; Text '丝'
   IOField "I/O 域_13" at 162,12 size 164x31; FormatPattern ????
      ProcessValue <- "数据变量.当前人员编号"
*)

(* ===== HMI "HMI_RT_1" =====

ScreenModuleEditorView "精炼机面板" 338x480
   Rectangle "备妥矩形" at 1,1 size 339x48
      Visibility <- "数据变量.开关量汇总"
   Rectangle "运行矩形" at 1,1 size 337x48
      Visibility <- "数据变量.开关量汇总"
   Rectangle "故障矩形" at 1,1 size 338x48
      Visibility <- "数据变量.开关量汇总"
   TextField "设备名称" at 8,11 size 107x28; Text 'N11号精炼机'
   IOField "I/O 域_1" at 8,72 size 154x80; FormatPattern 999
      ProcessValue <- "数据变量.滚筒电机电流"
   IOField "I/O 域_2" at 8,170 size 160x80; FormatPattern 99.9
      ProcessValue <- "数据变量.滚筒电机频率"
   TextField "文本域_2" at 118,218 size 28x26; Text 'HZ'
   TextField "文本域_3" at 118,132 size 17x26; Text 'A'
   TextField "文本域_4" at 9,49 size 37x26; Text '电流'
   TextField "文本域_5" at 9,148 size 37x26; Text '频率'
   IOField "I/O 域_3" at 186,69 size 120x80; FormatPattern 999
      ProcessValue <- "数据变量.滚筒电机功率"
   TextField "文本域_1" at 311,136 size 20x26; Text '%'
   TextField "文本域_6" at 200,46 size 37x26; Text '功率'
   IOField "I/O 域_4" at 187,171 size 104x80; FormatPattern 999
      ProcessValue <- "数据变量.胶温"
   TextField "文本域_7" at 309,218 size 21x26; Text '℃'
   TextField "文本域_8" at 203,149 size 37x26; Text '胶温'
   TextField "文本域_9" at 3,450 size 35x23; Text '计时:'
   TextField "文本域_10" at 158,450 size 35x23; Text '电能:'
   IOField "I/O 域_5" at 38,454 size 90x17; FormatPattern 9999999999
      ProcessValue <- "数据变量.滚筒电机计时"
   TextField "文本域_11" at 137,451 size 13x23; Text 'S'
   IOField "I/O 域_6" at 193,454 size 90x17; FormatPattern 9999999999
      ProcessValue <- "数据变量.滚筒电机电度"
   TextField "文本域_12" at 289,451 size 39x23; Text 'KWH'
   TextField "文本域_13" at 17,268 size 87x23; Text '左前滚筒轴温:'
   IOField "I/O 域_7" at 17,285 size 82x43; FormatPattern 999.9
      ProcessValue <- "数据变量.左前辊温度"
   TextField "文本域_14" at 109,297 size 18x23; Text '℃'
   TextField "文本域_15" at 204,268 size 87x23; Text '右前滚筒轴温:'
   IOField "I/O 域_8" at 201,284 size 82x43; FormatPattern 999.9
      ProcessValue <- "数据变量.右前辊温度"
   TextField "文本域_16" at 308,296 size 18x23; Text '℃'
   TextField "文本域_17" at 16,328 size 87x23; Text '左后滚筒轴温:'
   IOField "I/O 域_9" at 16,346 size 82x43; FormatPattern 999.9
      ProcessValue <- "数据变量.左后辊温度"
   TextField "文本域_18" at 108,357 size 18x23; Text '℃'
   TextField "文本域_19" at 204,329 size 87x23; Text '右后滚筒轴温:'
   IOField "I/O 域_10" at 201,345 size 82x43; FormatPattern 999.9
      ProcessValue <- "数据变量.右后辊温度"
   TextField "文本域_20" at 308,357 size 18x23; Text '℃'
   TextField "文本域_21" at 17,392 size 83x23; Text '左滚筒间隙值'
   IOField "I/O 域_11" at 12,408 size 82x43; FormatPattern 9999
      ProcessValue <- "数据变量.左间隙"
   TextField "文本域_22" at 109,421 size 18x23; Text '丝'
   TextField "文本域_23" at 205,393 size 87x23; Text '右滚筒间隙值:'
   IOField "I/O 域_12" at 200,408 size 82x43; FormatPattern 9999
      ProcessValue <- "数据变量.右间隙"
   TextField "文本域_24" at 309,420 size 18x23; Text '丝'
   IOField "I/O 域_13" at 162,12 size 164x31; FormatPattern ????
      ProcessValue <- "数据变量.当前人员编号"
*)

(* ===== HMI "HMI_RT_1" =====

ScreenModuleEditorView "精炼机面板" 338x480
   Rectangle "备妥矩形" at -1,12 size 339x48
      Visibility <- "数据变量.开关量汇总"
   Rectangle "运行矩形" at 1,24 size 337x48
      Visibility <- "数据变量.开关量汇总"
   Rectangle "故障矩形" at 0,60 size 338x48
      Visibility <- "数据变量.开关量汇总"
   TextField "设备名称" at 8,11 size 107x28; Text 'N11号精炼机'
   IOField "I/O 域_1" at 8,72 size 154x80; FormatPattern 999
      ProcessValue <- "数据变量.滚筒电机电流"
   IOField "I/O 域_2" at 8,170 size 160x80; FormatPattern 99.9
      ProcessValue <- "数据变量.滚筒电机频率"
   TextField "文本域_2" at 118,218 size 28x26; Text 'HZ'
   TextField "文本域_3" at 118,132 size 17x26; Text 'A'
   TextField "文本域_4" at 9,49 size 37x26; Text '电流'
   TextField "文本域_5" at 9,148 size 37x26; Text '频率'
   IOField "I/O 域_3" at 186,69 size 120x80; FormatPattern 999
      ProcessValue <- "数据变量.滚筒电机功率"
   TextField "文本域_1" at 311,136 size 20x26; Text '%'
   TextField "文本域_6" at 200,46 size 37x26; Text '功率'
   IOField "I/O 域_4" at 187,171 size 104x80; FormatPattern 999
      ProcessValue <- "数据变量.胶温"
   TextField "文本域_7" at 309,218 size 21x26; Text '℃'
   TextField "文本域_8" at 203,149 size 37x26; Text '胶温'
   TextField "文本域_9" at 3,450 size 35x23; Text '计时:'
   TextField "文本域_10" at 158,450 size 35x23; Text '电能:'
   IOField "I/O 域_5" at 38,454 size 90x17; FormatPattern 9999999999
      ProcessValue <- "数据变量.滚筒电机计时"
   TextField "文本域_11" at 137,451 size 13x23; Text 'S'
   IOField "I/O 域_6" at 193,454 size 90x17; FormatPattern 9999999999
      ProcessValue <- "数据变量.滚筒电机电度"
   TextField "文本域_12" at 289,451 size 39x23; Text 'KWH'
   TextField "文本域_13" at 17,268 size 87x23; Text '左前滚筒轴温:'
   IOField "I/O 域_7" at 17,285 size 82x43; FormatPattern 999.9
      ProcessValue <- "数据变量.左前辊温度"
   TextField "文本域_14" at 109,297 size 18x23; Text '℃'
   TextField "文本域_15" at 204,268 size 87x23; Text '右前滚筒轴温:'
   IOField "I/O 域_8" at 201,284 size 82x43; FormatPattern 999.9
      ProcessValue <- "数据变量.右前辊温度"
   TextField "文本域_16" at 308,296 size 18x23; Text '℃'
   TextField "文本域_17" at 16,328 size 87x23; Text '左后滚筒轴温:'
   IOField "I/O 域_9" at 16,346 size 82x43; FormatPattern 999.9
      ProcessValue <- "数据变量.左后辊温度"
   TextField "文本域_18" at 108,357 size 18x23; Text '℃'
   TextField "文本域_19" at 204,329 size 87x23; Text '右后滚筒轴温:'
   IOField "I/O 域_10" at 201,345 size 82x43; FormatPattern 999.9
      ProcessValue <- "数据变量.右后辊温度"
   TextField "文本域_20" at 308,357 size 18x23; Text '℃'
   TextField "文本域_21" at 17,392 size 83x23; Text '左滚筒间隙值'
   IOField "I/O 域_11" at 12,408 size 82x43; FormatPattern 9999
      ProcessValue <- "数据变量.左间隙"
   TextField "文本域_22" at 109,421 size 18x23; Text '丝'
   TextField "文本域_23" at 205,393 size 87x23; Text '右滚筒间隙值:'
   IOField "I/O 域_12" at 200,408 size 82x43; FormatPattern 9999
      ProcessValue <- "数据变量.右间隙"
   TextField "文本域_24" at 309,420 size 18x23; Text '丝'
   IOField "I/O 域_13" at 162,12 size 164x31; FormatPattern ????
      ProcessValue <- "数据变量.当前人员编号"
*)

(* ===== HMI "HMI_RT_1" =====

ScreenModuleEditorView "精炼机面板" 338x480
   Rectangle "备妥矩形" at 1,1 size 339x48
      Visibility <- "数据变量.开关量汇总"
   Rectangle "运行矩形" at 1,1 size 337x48
      Visibility <- "数据变量.开关量汇总"
   Rectangle "故障矩形" at 1,1 size 338x48
      Visibility <- "数据变量.开关量汇总"
   TextField "设备名称" at 8,11 size 107x28; Text 'N11号精炼机'
   IOField "I/O 域_1" at 8,72 size 154x80; FormatPattern 999
      ProcessValue <- "数据变量.滚筒电机电流"
   IOField "I/O 域_2" at 8,170 size 160x80; FormatPattern 99.9
      ProcessValue <- "数据变量.滚筒电机频率"
   TextField "文本域_2" at 118,218 size 28x26; Text 'HZ'
   TextField "文本域_3" at 118,132 size 17x26; Text 'A'
   TextField "文本域_4" at 9,49 size 37x26; Text '电流'
   TextField "文本域_5" at 9,148 size 37x26; Text '频率'
   IOField "I/O 域_3" at 186,69 size 120x80; FormatPattern 999
      ProcessValue <- "数据变量.滚筒电机功率"
   TextField "文本域_1" at 311,136 size 20x26; Text '%'
   TextField "文本域_6" at 200,46 size 37x26; Text '功率'
   IOField "I/O 域_4" at 187,171 size 104x80; FormatPattern 999
      ProcessValue <- "数据变量.胶温"
   TextField "文本域_7" at 309,218 size 21x26; Text '℃'
   TextField "文本域_8" at 203,149 size 37x26; Text '胶温'
   TextField "文本域_9" at 3,450 size 35x23; Text '计时:'
   TextField "文本域_10" at 158,450 size 35x23; Text '电能:'
   IOField "I/O 域_5" at 38,454 size 90x17; FormatPattern 9999999999
      ProcessValue <- "数据变量.滚筒电机计时"
   TextField "文本域_11" at 137,451 size 13x23; Text 'S'
   IOField "I/O 域_6" at 193,454 size 90x17; FormatPattern 9999999999
      ProcessValue <- "数据变量.滚筒电机电度"
   TextField "文本域_12" at 289,451 size 39x23; Text 'KWH'
   TextField "文本域_13" at 17,268 size 87x23; Text '左前滚筒轴温:'
   IOField "I/O 域_7" at 17,285 size 82x43; FormatPattern 999.9
      ProcessValue <- "数据变量.左前辊温度"
   TextField "文本域_14" at 109,297 size 18x23; Text '℃'
   TextField "文本域_15" at 204,268 size 87x23; Text '右前滚筒轴温:'
   IOField "I/O 域_8" at 201,284 size 82x43; FormatPattern 999.9
      ProcessValue <- "数据变量.右前辊温度"
   TextField "文本域_16" at 308,296 size 18x23; Text '℃'
   TextField "文本域_17" at 16,328 size 87x23; Text '左后滚筒轴温:'
   IOField "I/O 域_9" at 16,346 size 82x43; FormatPattern 999.9
      ProcessValue <- "数据变量.左后辊温度"
   TextField "文本域_18" at 108,357 size 18x23; Text '℃'
   TextField "文本域_19" at 204,329 size 87x23; Text '右后滚筒轴温:'
   IOField "I/O 域_10" at 201,345 size 82x43; FormatPattern 999.9
      ProcessValue <- "数据变量.右后辊温度"
   TextField "文本域_20" at 308,357 size 18x23; Text '℃'
   TextField "文本域_21" at 17,392 size 83x23; Text '左滚筒间隙值'
   IOField "I/O 域_11" at 12,408 size 82x43; FormatPattern 9999
      ProcessValue <- "数据变量.左间隙"
   TextField "文本域_22" at 109,421 size 18x23; Text '丝'
   TextField "文本域_23" at 205,393 size 87x23; Text '右滚筒间隙值:'
   IOField "I/O 域_12" at 200,408 size 82x43; FormatPattern 9999
      ProcessValue <- "数据变量.右间隙"
   TextField "文本域_24" at 309,420 size 18x23; Text '丝'
   IOField "I/O 域_13" at 162,12 size 164x31; FormatPattern ????
      ProcessValue <- "数据变量.当前人员编号"
*)